FUNCTION "RPA20B_Main" : Void   // FC43, SCL
{ S7_Optimized_Access := 'FALSE' }
VERSION : 0.1
BEGIN


       IF "RPA20B_manual_DOWN" THEN //manual move down
           "RPA20_motor_up" := false;
           "RPA20B_motor_down" := "RPA20B_manual_move";
       ELSIF "RPA20B_manual_UP" THEN // manual move up
           "RPA20_motor_up" := "RPA20B_manual_move";
           "RPA20B_motor_down" := false;
       ELSE // automatic mode operator 1
           "RPA20B_handler_op_1"();
       END_IF;

      "RPA20B_handler_op_2"();

      // blikání LED na tlačítkách

      "RPA20B_open_door_LED_green" := "Clock_0.5Hz" AND ("RPA20B_blend_presence_sensor_1" OR "RPA20B_blend_presence_sensor_2")AND (NOT "RPA20B_open_drawer");

      IF "RPA20B_datablock".RPA20B_station_monitoring_send = true THEN
          "RPA20B_datablock".RPA20B_station_monitoring_send := NOT "pa20b_station_monitoring"(station_activity_state := "RPA20B_ES_feedback",
                                                                                              blend_senzor_l := "RPA20B_blend_presence_sensor_2",
                                                                                              blend_senzor_r := "RPA20B_blend_presence_sensor_1",
                                                                                              server_connection := "tcp_datablock".tcp_connection,
                                                                                              index:="tcp_datablock".<??.?>);
      ELSE
          IF "RPA20B_datablock".RPA20B_activity_state_pre <> "RPA20B_ES_feedback" OR 
              "RPA20B_datablock".RPA20B_left_cover_pressence_sensor_pre <> "RPA20B_blend_presence_sensor_2" OR
              "RPA20B_datablock".RPA20B_right_cover_pressence_sensor_pre <> "RPA20B_blend_presence_sensor_1" THEN
              "RPA20B_datablock".RPA20B_station_monitoring_send := true;
          END_IF;

          "RPA20B_datablock".RPA20B_activity_state_pre := "RPA20B_ES_feedback";
          "RPA20B_datablock".RPA20B_left_cover_pressence_sensor_pre := "RPA20B_blend_presence_sensor_2";
          "RPA20B_datablock".RPA20B_right_cover_pressence_sensor_pre := "RPA20B_blend_presence_sensor_1";
      END_IF;
      IF "RPA20B_manual_UP" THEN
          "RPA20B_Camera_Result_OK" := false;
          "RPA20B_Camera_Result_NOK" := false;
      END_IF;
      "RPA20B_Camera_Trigger" := "RPA20B_Camera_Start_Test";
      "RPA20B_Camera_TrafficLight_Green" := "RPA20B_Camera_Result_OK";
      "RPA20B_Camera_TrafficLight_Red" := "RPA20B_Camera_Result_NOK";
END_FUNCTION

FUNCTION "build_new_record" : Void   // FC44, SCL
{ S7_Optimized_Access := 'FALSE' }
VERSION : 0.1
BEGIN


   #temp_string := CONCAT(IN1 := '$'172', IN2 := "RPA60_DataBlock".RPA60_frame_order);
   #temp_string := CONCAT(IN1 := #temp_string, IN2 := '$', ');
   Strg_TO_Chars(Strg := #temp_string,
                 pChars := 0,
                 Cnt => #i,
                 Chars := #temp_record);

   #chars := 0;
   WHILE #record_in[#chars] <> '?' DO
       #temp_record[#chars+#i] := #record_in[#chars];
      #chars := #chars + 1;
   END_WHILE;

   #temp_record[#chars + #i] := '$L';
   #record_data := #temp_record;

   #i := 0;
   Strg_TO_Chars(Strg:='$'ID$' ,$'frame_code$', $'frame_order$', $'configuration$', $'PA30R_date_time$', $'PA60R_date_time$', ',
                 pChars:=0,
                 Cnt=>#chars,
                 Chars:=#temp_record);

   Strg_TO_Chars(Strg := '$'PA30R_Primer_207_SIKA$', $'PA30R_Remover_208_SIKA$', $'PA30R_rework$', $'PA60R_rework$', $'PA30R_cyclus_completed$', $'PA60R_cyclus_completed$'$L',
                 pChars := #chars,
                 Cnt => #i,
                 Chars := #temp_record);

   #record_items := #temp_record;
END_FUNCTION

FUNCTION "copyAndFill" : Void   // FC45, SCL
{ S7_Optimized_Access := 'FALSE' }
VERSION : 0.1
BEGIN




   //copy the input string to the output string
   #index := 1;
   #inputStringLen := LEN(#stringIn);
   #copyAndFill := '';
   IF #char_number >= #inputStringLen THEN
       WHILE #index <= #char_number DO
           IF #index >= (#char_number - #inputStringLen+1) THEN
               IF #stringIn[#index - (#char_number - #inputStringLen)] <> #charReplace THEN
                   #copyAndFill := CONCAT(IN1 := #copyAndFill, IN2 := #stringIn[#index - (#char_number - #inputStringLen)]);
               ELSE
                   #copyAndFill := CONCAT(IN1 := #copyAndFill, IN2 := #characterFill);
               END_IF;
           ELSE
               #copyAndFill := CONCAT(IN1 := #copyAndFill, IN2 := #characterFill);
           END_IF;

           #index := #index + 1;
       END_WHILE;
   END_IF;
END_FUNCTION

FUNCTION "RPA10B_handler_function" : Void   // FC48, SCL
{ S7_Optimized_Access := 'FALSE' }
VERSION : 0.1
BEGIN
END_FUNCTION

FUNCTION "RPA10B_idler_presence_handler" : Void   // FC49, SCL
{ S7_Optimized_Access := 'FALSE' }
VERSION : 0.1
BEGIN

   (*
   pokud je big fail state odemčený pak se podprogram vykoná

   pokud přítlačné kolečko ve stavu využíváno pak je rozlišováno jestli se jedná o stav ve kterém se čeká na vyjmutí z dokovací stanice a nebo jestli již je vyjmuto z dokovací stanice

   pokud se jedná o stav kdy se čeká na vyjmutí z dokovací stanice musí blikat světelná kontrolka přítlačného kolečka a být nastaven vnitřní stav stanice OK

   pokud se jedná o stav kdy již je přítlačné kolečko z dokovací stanice vyjmuto kontroluje se zda není vloženo zpátky před expirací časovače

   pokud je přítlačné kolečko vloženo do dokovací stanice před expirací časovače dojde k nastavení stavu big fail a blikání světelné kontrolky přítlačného kolečka

   *)

   IF (#bigFailStateLock = 0 OR #bigFailStateLock = #bigFailStateIdentifire OR #bigFailStateLock = #bigFailStateIdentifire + 100) AND
       #errorStateLock = 0 AND
       #fatalErrorStateLock = 0 THEN

       //blikání a svícení světelné kontrolky přítlačného kolečka
       //#bottlePresenceSensor AND "Clock_0.5Hz" AND #bottleInUsage
      // #rollerLED := (NOT #rollerPresenceSensor) OR (#rollerPresenceSensor AND "Clock_0.5Hz" AND #roller_in_use);
       //#rollerLED := (NOT #rollerPresenceSensor) OR (#rollerPresenceSensor AND #rollerUsageInterval[#workCyclusControlVariable] AND "Clock_0.5Hz");

       IF #bigFailStateLock = #bigFailStateIdentifire  THEN
           "setOKState"(confirm := true,
                        identifier := #bigFailStateIdentifire,
                        confirm_blinking := false,
                        blinkConfirmButton => #confirmButtonLed,
                        stateLock := #bigFailStateLock);
       ELSIF #bigFailStateLock = #bigFailStateIdentifire+100 AND #idler_presence_sensor = true THEN
               "setOKState"(confirm := #confirmButton,
                            identifier := #bigFailStateIdentifire+100,
                            confirm_blinking := true,
                            blinkConfirmButton => #confirmButtonLed,
                            stateLock := #bigFailStateLock);
       END_IF;
       //kontrola přítomnosti kolečka v pracovním cyklu
       IF #idler_in_use THEN
           "RPA10B_datablock".RPA10B_idler_checking_dalay := false;
           //nekontroluje první stav a poslední stav ve kterém je přítlačné kolečko používáno -> stav ve kterém se mění mění přítomnost kolečka v dokovací stanici
               IF #idler_presence_sensor THEN
                   IF #idler_taking THEN
                       IF "setBigFailState"(identifier := #bigFailStateIdentifire,
                                                error_state_lock:="RPA10B_datablock".PA10B_error_state_lock, fatal_state_error:="RPA10B_datablock".PA10B_fatal_error_state_lock, badfailStateLock := #bigFailStateLock) THEN
                           ;
                       END_IF;
                   END_IF;
               END_IF;
        ELSE
            IF (NOT #idler_presence_sensor) THEN
                IF "RPA10B_datablock".RPA10B_idler_checking_dalay THEN
                    IF "setBigFailState"(identifier := #bigFailStateIdentifire + 100,
                                             error_state_lock := "RPA10B_datablock".PA10B_error_state_lock, fatal_state_error := "RPA10B_datablock".PA10B_fatal_error_state_lock, badfailStateLock := #bigFailStateLock) THEN
                        ;
                    END_IF;
                ELSE
                    "RPA10B_datablock".RPA10B_idler_checking_dalay := "Clock_0.5Hz";
                END_IF;
            END_IF;
       END_IF;
   END_IF;
END_FUNCTION

FUNCTION "server_connection_handler" : Void   // FC50, SCL
{ S7_Optimized_Access := 'FALSE' }
VERSION : 0.1
BEGIN
   IF #database_connection = true THEN
       IF #error_state_lock = #error_state_lock_identifier THEN
           #error_state_lock := 0;
       END_IF;
   ELSE
       IF #fatal_error_state_lock = 0 AND #error_state_lock = 0 THEN
           #error_state_lock := #error_state_lock_identifier;
       END_IF;
   END_IF;
END_FUNCTION

FUNCTION "station_reset" : Void   // FC51, SCL
{ S7_Optimized_Access := 'FALSE' }
VERSION : 0.1
BEGIN
   #index := 1;

   WHILE (#index < 6) DO
       #fs_funel_control[#index] := false;
       #fs_show_fill_button[#index] := false;
       #index := #index + 1;
   END_WHILE;

   #funel_1 := false;
   #funel_2 := false;
   #funel_3 := false;
   #funel_4 := false;
   #funel_5 := false;

   #fs_chemical_type := 0;
   #hmi_label_index := 0;


   #fill_bottle_step := 9;
   #shake_deinit := true;
   #print_sp_bottle_label_step := 8;



   #fs_show_manual_or_scan := false;
   #fs_show_button := false;
   #fs_reset_e := false;
END_FUNCTION

FUNCTION "time_compare" : Void   // FC52, LAD
{ S7_Optimized_Access := 'FALSE' }
VERSION : 0.1
BEGIN

REGION Network 1
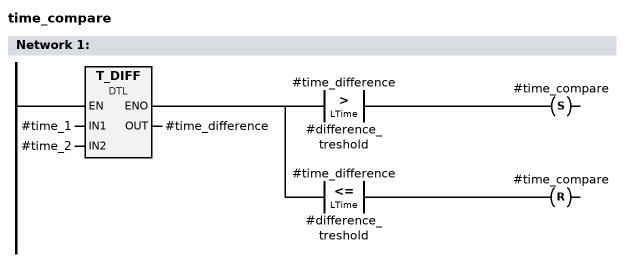
   // ENO of a box is taken as its EN; it also drops when the box reports an error
   #time_difference := T_DIFF(IN1 := #time_1, IN2 := #time_2);
   IF #time_difference > #difference_treshold THEN #time_compare := TRUE; END_IF;
   IF #time_difference <= #difference_treshold THEN #time_compare := FALSE; END_IF;
END_REGION
END_FUNCTION

FUNCTION "RPA30_Handler_function_A" : Void   // FC53, SCL
{ S7_Optimized_Access := 'FALSE' }
VERSION : 0.1
BEGIN
END_FUNCTION

FUNCTION "pa10r_station_monitoring" : Void   // FC54, SCL
{ S7_Optimized_Access := 'FALSE' }
VERSION : 0.1
BEGIN
   #pa10r_station_monitoring := false;
   (*
   IF #server_connection = true THEN
       IF "send_msg_to_pc_DB".DONE THEN
           "rcv_msg_from_pc_DB"(size := 1024,
                                time_out_interval := #lock);

           IF "rcv_msg_from_pc_DB".time_out = true THEN
               "send_msg_to_pc_DB".DONE := false;
               "rcv_msg_from_pc_DB".DONE := false;
               #server_connection := false;
           END_IF;

           IF "rcv_msg_from_pc_DB".DONE THEN
               "send_msg_to_pc_DB".DONE := false;
               "rcv_msg_from_pc_DB".DONE := false;
               "send_msg_to_pc_DB".synchronization := 0;
               "rcv_msg_from_pc_DB".synchronization := 0;
               #server_connection := true;
               #pa10r_station_monitoring := true;
           END_IF;
       ELSE

           //command 
           Strg_TO_Chars(Strg := 'PA10R_STATE~',
                         pChars := 0,
                         Cnt => #chars,
                         Chars := #chars_out);
           #i := #chars;

           // station state 
           IF #station_activity_state = true THEN
               IF #fatal_error_state > 0 THEN
                   CASE #fatal_error_state OF
                       150:
                           Strg_TO_Chars(Strg := '<html>Station state: Y axis<br>valve lock error</html>~',
                                         pChars := #i,
                                         Cnt => #chars,
                                         Chars := #chars_out);
                       160:
                           Strg_TO_Chars(Strg := '<html>Station state: X axis<br>valve lock error</html>~',
                                         pChars := #i,
                                         Cnt => #chars,
                                         Chars := #chars_out);
                       ELSE
                           Strg_TO_Chars(Strg := 'Station state: Unknown~',
                                         pChars := #i,
                                         Cnt => #chars,
                                         Chars := #chars_out);
                   END_CASE;
               ELSE
                   IF #error_state > 0 THEN
                       Strg_TO_Chars(Strg := 'Station state: Unknown~',
                                     pChars := #i,
                                     Cnt => #chars,
                                     Chars := #chars_out);
                   ELSE
                       IF #big_fail_state > 0 THEN
                           Strg_TO_Chars(Strg := 'Station state: Unknown~',
                                         pChars := #i,
                                         Cnt => #chars,
                                         Chars := #chars_out);
                       ELSE
                           IF #fail_state > 0 THEN
                               CASE #fail_state OF
                                   110:
                                       Strg_TO_Chars(Strg := 'Station state: Felt box is empty~',
                                                     pChars := #i,
                                                     Cnt => #chars,
                                                     Chars := #chars_out);
                                   200:  // Statement section case 2 to 4
                                       Strg_TO_Chars(Strg := '<html>Station state: Primer DV594V1<br>in primer box</html>~',
                                                     pChars := #i,
                                                     Cnt => #chars,
                                                     Chars := #chars_out);
                                   201:
                                       Strg_TO_Chars(Strg := '<html>Station state: Activator DW646<br>in primer box</html>~',
                                                     pChars := #i,
                                                     Cnt => #chars,
                                                     Chars := #chars_out);
                                   202:
                                       Strg_TO_Chars(Strg := '<html>Station state: Primer 207<br>in primer box</html>~',
                                                     pChars := #i,
                                                     Cnt => #chars,
                                                     Chars := #chars_out);
                                   300:
                                       Strg_TO_Chars(Strg := '<html>Station state: Primer DV594V1<br>out of primer box</html>~',
                                                     pChars := #i,
                                                     Cnt => #chars,
                                                     Chars := #chars_out);
                                   301:
                                       Strg_TO_Chars(Strg := '<html>Station state: Activator DW646<br>out of primer box</html>~',
                                                     pChars := #i,
                                                     Cnt => #chars,
                                                     Chars := #chars_out);
                                   302:
                                       Strg_TO_Chars(Strg := '<html>Station state: Primer 207<br>out of primer box</html>~',
                                                     pChars := #i,
                                                     Cnt => #chars,
                                                     Chars := #chars_out);
                                   303:
                                       Strg_TO_Chars(Strg := '<html>Station state: Remover 208<br>out of primer box</html>~',
                                                     pChars := #i,
                                                     Cnt => #chars,
                                                     Chars := #chars_out);
                                   6:
                                       Strg_TO_Chars(Strg := 'Station state: Remover 208 expired~',
                                                     pChars := #i,
                                                     Cnt => #chars,
                                                     Chars := #chars_out);
                                   ELSE  // Statement section ELSE
                                       Strg_TO_Chars(Strg := 'Station state: Unknown~',
                                                     pChars := #i,
                                                     Cnt => #chars,
                                                     Chars := #chars_out);
                               END_CASE;

                           ELSE
                               Strg_TO_Chars(Strg := 'Station state: OK~',
                                             pChars := #i,
                                             Cnt => #chars,
                                             Chars := #chars_out);
                           END_IF;
                       END_IF;
                   END_IF;
               END_IF;
           ELSE
               Strg_TO_Chars(Strg := 'Station state: Inactive~',
                             pChars := #i,
                             Cnt => #chars,
                             Chars := #chars_out);
           END_IF;

           #i := #i+#chars;

           // work cyclus state 

           IF #work_cyclus_state = "RPA10R_hmi_go_to_home_position" THEN
               Strg_TO_Chars(Strg := 'Work cyclus state: Waiting for home position~',
                             pChars := #i,
                             Cnt => #chars,
                             Chars := #chars_out);
           ELSIF #work_cyclus_state = "RPA10R_hmi_scan_frame" THEN
               Strg_TO_Chars(Strg := 'Work cyclus state: Scan frame~',
                             pChars := #i,
                             Cnt => #chars,
                             Chars := #chars_out);
           ELSIF #work_cyclus_state = "RPA10R_hmi_take_bottle_1" THEN
               Strg_TO_Chars(Strg := 'Work cyclus state: Take activator DW 646~',
                             pChars := #i,
                             Cnt => #chars,
                             Chars := #chars_out);
           ELSIF #work_cyclus_state = "RPA10R_hmi_scan_bottle" THEN
               Strg_TO_Chars(Strg := 'Work cyclus state: Scan bottle~',
                             pChars := #i,
                             Cnt => #chars,
                             Chars := #chars_out);
           ELSIF #work_cyclus_state = "RPA10R_hmi_change_pad" THEN
               Strg_TO_Chars(Strg := 'Work cyclus state: Change pad~',
                             pChars := #i,
                             Cnt => #chars,
                             Chars := #chars_out);
           ELSIF #work_cyclus_state = "RPA10R_hmi_apply_bottle_1_on_side_5_5" OR #work_cyclus_state = "RPA10R_hmi_apply_bottle_1_on_side_5" THEN
               Strg_TO_Chars(Strg := 'Work cyclus state: Apply activator on frame~',
                             pChars := #i,
                             Cnt => #chars,
                             Chars := #chars_out);
           ELSIF #work_cyclus_state = "RPA10R_hmi_turn_clockwise" THEN
               Strg_TO_Chars(Strg := 'Work cyclus state: Turn frame clockwise~',
                             pChars := #i,
                             Cnt => #chars,
                             Chars := #chars_out);
           ELSIF #work_cyclus_state = "RPA10R_hmi_take_bottle_2" THEN
               Strg_TO_Chars(Strg := 'Work cyclus state: Take bottle of primer DV954~',
                             pChars := #i,
                             Cnt => #chars,
                             Chars := #chars_out);
           ELSIF #work_cyclus_state = "RPA10R_hmi_whipe_off_side_5_5" OR #work_cyclus_state = "RPA10R_hmi_whipe_off_side_5" THEN
               Strg_TO_Chars(Strg := '<html>Work cyclus state: Wipe off activator<br> from frame</html>~',
                             pChars := #i,
                             Cnt => #chars,
                             Chars := #chars_out);
           ELSIF #work_cyclus_state = "RPA10R_hmi_apply_bottle_2_on_side_5_5" OR #work_cyclus_state = "RPA10R_hmi_apply_bottle_2_on_side_5" THEN
               Strg_TO_Chars(Strg := 'Work cyclus state: Apply primer on frame~',
                             pChars := #i,
                             Cnt => #chars,
                             Chars := #chars_out);
           ELSIF #work_cyclus_state = "RPA10R_hmi_put_back_bottle_1" THEN
               Strg_TO_Chars(Strg := '<html>Work cyclus state: Put activator DW 646<br>bottle to primer bar</html>~',
                             pChars := #i,
                             Cnt => #chars,
                             Chars := #chars_out);
           ELSIF #work_cyclus_state = "RPA10R_hmi_put_back_bottle_2" THEN
               Strg_TO_Chars(Strg := '<html>Work cyclus state: Put primer DV954 bottle<br>to primer bar</html>~',
                             pChars := #i,
                             Cnt => #chars,
                             Chars := #chars_out);
           ELSIF #work_cyclus_state = "RPA10R_hmi_take_felt" THEN
               Strg_TO_Chars(Strg := 'Work cyclus state: Take felt~',
                             pChars := #i,
                             Cnt => #chars,
                             Chars := #chars_out);
           ELSIF #work_cyclus_state = "RPA10R_hmi_turn_horizontaly" THEN
               Strg_TO_Chars(Strg := 'Work cyclus state: Turn frame horizontaly~',
                             pChars := #i,
                             Cnt => #chars,
                             Chars := #chars_out);
           ELSIF #work_cyclus_state = "RPA10R_hmi_on_felt_apply_remover" THEN
               Strg_TO_Chars(Strg := 'Work cyclus state: On felt apply remover~',
                             pChars := #i,
                             Cnt => #chars,
                             Chars := #chars_out);
           ELSIF #work_cyclus_state = "RPA10R_hmi_apply_remover_to_side_5" THEN
               Strg_TO_Chars(Strg := 'Work cyclus state: Apply remover 208 on frame~',
                             pChars := #i,
                             Cnt => #chars,
                             Chars := #chars_out);
           ELSIF #work_cyclus_state = "RPA10R_hmi_turn_counterclockwise" THEN
               Strg_TO_Chars(Strg := 'Work cyclus state: Turn frame counterclockwise~',
                             pChars := #i,
                             Cnt => #chars,
                             Chars := #chars_out);
           ELSIF #work_cyclus_state = "RPA10R_hmi_take_bottle_3" THEN
               Strg_TO_Chars(Strg := 'Work cyclus state: Take bottle of primer 207~',
                             pChars := #i,
                             Cnt => #chars,
                             Chars := #chars_out);
           ELSIF #work_cyclus_state = "RPA10R_hmi_put_back_bottle_3" THEN
               Strg_TO_Chars(Strg := '<html>Work cyclus state: Put primer 207 bottle <br> to primer bar</html>~',
                             pChars := #i,
                             Cnt => #chars,
                             Chars := #chars_out);
           ELSIF #work_cyclus_state = "RPA10R_hmi_end_of_cyclus" THEN
               Strg_TO_Chars(Strg := 'Work cyclus state: End of work cyclus~',
                             pChars := #i,
                             Cnt => #chars,
                             Chars := #chars_out);
           ELSIF #work_cyclus_state = 254 THEN
               Strg_TO_Chars(Strg := 'Work cyclus state: Manual mode~',
                             pChars := #i,
                             Cnt => #chars,
                             Chars := #chars_out);
           ELSE
               Strg_TO_Chars(Strg := 'Work cyclus state: Unknown~',
                             pChars := #i,
                             Cnt => #chars,
                             Chars := #chars_out);
           END_IF;

           #i := #i+#chars;
           // home position 
           IF #position_sensor_y AND #position_sensor_x THEN
               Strg_TO_Chars(Strg := 'Home position: Yes~',
                             pChars := #i,
                             Cnt => #chars,
                             Chars := #chars_out);
           ELSE
               Strg_TO_Chars(Strg := 'Home position: No~',
                             pChars := #i,
                             Cnt => #chars,
                             Chars := #chars_out);
           END_IF;

           #i := #i + #chars;
           // current frame code
           Strg_TO_Chars(Strg := 'Current frame code: ',
                         pChars := #i,
                         Cnt => #chars,
                         Chars := #chars_out);
           #i := #i + #chars;
           IF #current_frame_code <> '' THEN
               Strg_TO_Chars(Strg := #current_frame_code,
                             pChars := #i,
                             Cnt => #chars,
                             Chars := #chars_out);
           ELSE
               Strg_TO_Chars(Strg := 'None',
                             pChars := #i,
                             Cnt => #chars,
                             Chars := #chars_out);
           END_IF;
           #i := #i + #chars;

           // station configuration
           IF #station_configuration = 0 THEN
               Strg_TO_Chars(Strg := '~Station configuration: 581A~',
                             pChars := #i,
                             Cnt => #chars,
                             Chars := #chars_out);
           ELSIF #station_configuration = 1 THEN
               Strg_TO_Chars(Strg := '~Station configuration: 581B~',
                             pChars := #i,
                             Cnt => #chars,
                             Chars := #chars_out);
           ELSIF #station_configuration = 2 THEN
               Strg_TO_Chars(Strg := '~Station configuration: 582A~',
                             pChars := #i,
                             Cnt => #chars,
                             Chars := #chars_out);
           ELSIF #station_configuration = 3 THEN
               Strg_TO_Chars(Strg := '~Station configuration: 582B~',
                             pChars := #i,
                             Cnt => #chars,
                             Chars := #chars_out);
           END_IF;

           #i := #i + #chars;

           "send_msg_to_pc_DB"(lock := #chars_out,
                               lock := 1024,
                               time_out_interval := #i,
                               time_out_interval := #lock);
           IF "send_msg_to_pc_DB".time_out = true THEN
               #server_connection := false;
           END_IF;
       END_IF;
   END_IF;
   *)
END_FUNCTION

FUNCTION "pa50r_station_monitoring" : Void   // FC55, SCL
{ S7_Optimized_Access := 'FALSE' }
VERSION : 0.1
BEGIN
   #pa50r_station_monitoring := false;
   (*
   IF #server_connection = true THEN
       IF "send_msg_to_pc_DB".DONE THEN
           "rcv_msg_from_pc_DB"(size := 1024,
                                time_out_interval := #lock);

           IF "rcv_msg_from_pc_DB".time_out = true THEN
               "send_msg_to_pc_DB".DONE := false;
               "rcv_msg_from_pc_DB".DONE := false;
               #server_connection := false;
           END_IF;

           IF "rcv_msg_from_pc_DB".DONE THEN
               "send_msg_to_pc_DB".DONE := false;
               "rcv_msg_from_pc_DB".DONE := false;
               "send_msg_to_pc_DB".synchronization := 0;
               "rcv_msg_from_pc_DB".synchronization := 0;
               #server_connection := true;
               #pa50r_station_monitoring := true;
           END_IF;
       ELSE

           //command 
           Strg_TO_Chars(Strg := 'PA50R_STATE~',
                         pChars := 0,
                         Cnt => #chars,
                         Chars := #chars_out);
           #i := #chars;

           //station state
           IF #station_activity_state = true THEN
               IF #fatal_error_state > 0 THEN
                   Strg_TO_Chars(Strg := 'Station state: Unknown~',
                                 pChars := #i,
                                 Cnt => #chars,
                                 Chars := #chars_out);
               ELSE
                   IF #error_state > 0 THEN
                       CASE #error_state OF
                           21000:
                               Strg_TO_Chars(Strg := 'Station state: Frame already processed~',
                                             pChars := #i,
                                             Cnt => #chars,
                                             Chars := #chars_out);
                           22000:
                               Strg_TO_Chars(Strg := 'Station state:Frame was not on previous station~',
                                             pChars := #i,
                                             Cnt => #chars,
                                             Chars := #chars_out);
                           23000:
                               Strg_TO_Chars(Strg := 'Station state: Frame has more then 8 hours~',
                                             pChars := #i,
                                             Cnt => #chars,
                                             Chars := #chars_out);
                           24000:
                               Strg_TO_Chars(Strg := 'Station state: Frame has less then 10 minutes~',
                                             pChars := #i,
                                             Cnt => #chars,
                                             Chars := #chars_out);
                           25000:
                               Strg_TO_Chars(Strg := 'Station state: Frame is not in database~',
                                             pChars := #i,
                                             Cnt => #chars,
                                             Chars := #chars_out);
                           26000:
                               Strg_TO_Chars(Strg := 'Station state: Bad station configuration~',
                                             pChars := #i,
                                             Cnt => #chars,
                                             Chars := #chars_out);
                           ELSE  // Statement section ELSE
                               Strg_TO_Chars(Strg := 'Station state: Unknown~',
                                             pChars := #i,
                                             Cnt => #chars,
                                             Chars := #chars_out);
                       END_CASE;

                       Strg_TO_Chars(Strg := 'Station state: Unknown~',
                                     pChars := #i,
                                     Cnt => #chars,
                                     Chars := #chars_out);
                   ELSE
                       IF #big_fail_state > 0 THEN
                           Strg_TO_Chars(Strg := 'Station state: Unknown~',
                                         pChars := #i,
                                         Cnt => #chars,
                                         Chars := #chars_out);
                       ELSE
                           IF #fail_state > 0 THEN
                                       Strg_TO_Chars(Strg := 'Station state: Unknown~',
                                                     pChars := #i,
                                                     Cnt => #chars,
                                                     Chars := #chars_out);
                           ELSE
                               Strg_TO_Chars(Strg := 'Station state: OK~',
                                             pChars := #i,
                                             Cnt => #chars,
                                             Chars := #chars_out);
                           END_IF;
                       END_IF;
                   END_IF;
               END_IF;
           ELSE
               Strg_TO_Chars(Strg := 'Station state: Inactive~',
                             pChars := #i,
                             Cnt => #chars,
                             Chars := #chars_out);
           END_IF;

           #i := #i+#chars;

           //work cyclus state

           IF #work_cyclus_state = "RPA50_hmi_go_to_home_position" THEN
               Strg_TO_Chars(Strg := 'Work cyclus state: Waiting for home position~',
                             pChars := #i,
                             Cnt => #chars,
                             Chars := #chars_out);
           ELSIF #work_cyclus_state = "RPA50_hmi_scan_frame" THEN
               Strg_TO_Chars(Strg := 'Work cyclus state: Scan frame code~',
                             pChars := #i,
                             Cnt => #chars,
                             Chars := #chars_out);
           ELSIF #work_cyclus_state = "RPA50_hmi_apply_tape" THEN
               Strg_TO_Chars(Strg := '<html>Work cyclus state: Application of tape <br>on every sides of grame</hmt>~',
                             pChars := #i,
                             Cnt => #chars,
                             Chars := #chars_out);
           ELSIF #work_cyclus_state = "RPA50_hmi_end_of_cyclus" THEN
               Strg_TO_Chars(Strg := 'Work cyclus state: End of work cyclus~',
                             pChars := #i,
                             Cnt => #chars,
                             Chars := #chars_out);
           ELSE
               Strg_TO_Chars(Strg := 'Work cyclus state: Unknown~',
                             pChars := #i,
                             Cnt => #chars,
                             Chars := #chars_out);
           END_IF;

           #i := #i+#chars;
           //home position
           IF #position_sensor_y THEN
               Strg_TO_Chars(Strg := 'Home position: Yes~',
                             pChars := #i,
                             Cnt => #chars,
                             Chars := #chars_out);
           ELSE
               Strg_TO_Chars(Strg := 'Home position: No~',
                             pChars := #i,
                             Cnt => #chars,
                             Chars := #chars_out);
           END_IF;

           #i := #i + #chars;
           //current frame code
           Strg_TO_Chars(Strg := 'Current frame code: ',
                         pChars := #i,
                         Cnt => #chars,
                         Chars := #chars_out);
           #i := #i + #chars;
           IF #current_frame_code <> '' THEN
               Strg_TO_Chars(Strg := #current_frame_code,
                             pChars := #i,
                             Cnt => #chars,
                             Chars := #chars_out);
           ELSE
               Strg_TO_Chars(Strg := 'None',
                             pChars := #i,
                             Cnt => #chars,
                             Chars := #chars_out);
           END_IF;
           #i := #i + #chars;

           //station configuration
           IF #station_configuration = 0 THEN
               Strg_TO_Chars(Strg := '~Station configuration: 581A',
                             pChars := #i,
                             Cnt => #chars,
                             Chars := #chars_out);
           ELSIF #station_configuration = 1 THEN
               Strg_TO_Chars(Strg := '~Station configuration: 581B',
                             pChars := #i,
                             Cnt => #chars,
                             Chars := #chars_out);
           ELSIF #station_configuration = 2 THEN
               Strg_TO_Chars(Strg := '~Station configuration: 582A',
                             pChars := #i,
                             Cnt => #chars,
                             Chars := #chars_out);
           ELSIF #station_configuration = 3 THEN
               Strg_TO_Chars(Strg := '~Station configuration: 582B',
                             pChars := #i,
                             Cnt => #chars,
                             Chars := #chars_out);
           END_IF;

           #i := #i + #chars;

           "send_msg_to_pc_DB"(time_out_interval := #chars_out,
                               time_out_interval := 1024,
                               lock := #i,
                               lock := #lock);
           IF "send_msg_to_pc_DB".time_out = true THEN
               #server_connection := false;
           END_IF;
       END_IF;
   END_IF;
   *)
END_FUNCTION

FUNCTION "pa60r_station_monitoring" : Void   // FC56, SCL
{ S7_Optimized_Access := 'FALSE' }
VERSION : 0.1
BEGIN
   #pa60r_station_monitoring := false;
   IF #server_connection = true THEN
       IF #index = 255 THEN
       (* command *)
           Strg_TO_Chars(Strg := 'PA60R_STATE~',
                         pChars := 0,
                         Cnt => #chars,
                         Chars := #temp_buffer);
           #i := #chars;

           (* station state *)
           IF #station_activity_state = true THEN
               IF #fatal_error_state > 0 THEN
                   CASE #fatal_error_state OF
                       150:  // Statement section case 1
                           Strg_TO_Chars(Strg := 'Station state: Y axis valve lock error~',
                                         pChars := #i,
                                         Cnt => #chars,
                                         Chars := #temp_buffer);
                       170:
                           Strg_TO_Chars(Strg := 'Station state: Bad frame code~',
                                         pChars := #i,
                                         Cnt => #chars,
                                         Chars := #temp_buffer);
                       180:
                           Strg_TO_Chars(Strg := 'Station state: Bad hardware configuration~',
                                         pChars := #i,
                                         Cnt => #chars,
                                         Chars := #temp_buffer);
                       230:
                           Strg_TO_Chars(Strg := 'Station state: Seal presence error~',
                                         pChars := #i,
                                         Cnt => #chars,
                                         Chars := #temp_buffer);
                       293:
                           Strg_TO_Chars(Strg := 'Station state: Change sealing fixtures~',
                                         pChars := #i,
                                         Cnt => #chars,
                                         Chars := #temp_buffer);
                       ELSE  // Statement section ELSE
                           Strg_TO_Chars(Strg := 'Station state: Unknown~',
                                         pChars := #i,
                                         Cnt => #chars,
                                         Chars := #temp_buffer);
                   END_CASE;
               ELSE
                   IF #error_state > 0 THEN
                       CASE #error_state OF
                           20000:
                               Strg_TO_Chars(Strg := 'Station state: Frame already processed~',
                                             pChars := #i,
                                             Cnt => #chars,
                                             Chars := #temp_buffer);
                           21000:
                               Strg_TO_Chars(Strg := 'Station state:Frame was not on previous station~',
                                             pChars := #i,
                                             Cnt => #chars,
                                             Chars := #temp_buffer);
                           23000:
                               Strg_TO_Chars(Strg := 'Station state: Frame has more then 8 hours~',
                                             pChars := #i,
                                             Cnt => #chars,
                                             Chars := #temp_buffer);
                           24000:
                               Strg_TO_Chars(Strg := 'Station state: Frame has less then 10 minutes~',
                                             pChars := #i,
                                             Cnt => #chars,
                                             Chars := #temp_buffer);
                           25000:
                               Strg_TO_Chars(Strg := 'Station state: Frame is not in database~',
                                             pChars := #i,
                                             Cnt => #chars,
                                             Chars := #temp_buffer);
                           26000:
                               Strg_TO_Chars(Strg := 'Station state: Bad station configuration~',
                                             pChars := #i,
                                             Cnt => #chars,
                                             Chars := #temp_buffer);
                           ELSE  // Statement section ELSE
                               Strg_TO_Chars(Strg := 'Station state: Unknown~',
                                             pChars := #i,
                                             Cnt => #chars,
                                             Chars := #temp_buffer);
                       END_CASE;

                       Strg_TO_Chars(Strg := 'Station state: Unknown~',
                                     pChars := #i,
                                     Cnt => #chars,
                                     Chars := #temp_buffer);
                   ELSE
                       IF #big_fail_state > 0 THEN
                           CASE #big_fail_state OF
                               120:  // Statement section case 1
                                   Strg_TO_Chars(Strg := 'Station state: Roller out of home position~',
                                                 pChars := #i,
                                                 Cnt => #chars,
                                                 Chars := #temp_buffer);

                               ELSE
                                   Strg_TO_Chars(Strg := 'Station state: Unknown~',
                                                 pChars := #i,
                                                 Cnt => #chars,
                                                 Chars := #temp_buffer);
                           END_CASE;


                       ELSE
                           IF #fail_state > 0 THEN
                               Strg_TO_Chars(Strg := 'Station state: Unknown~',
                                             pChars := #i,
                                             Cnt => #chars,
                                             Chars := #temp_buffer);
                           ELSE
                               Strg_TO_Chars(Strg := 'Station state: OK~',
                                             pChars := #i,
                                             Cnt => #chars,
                                             Chars := #temp_buffer);
                           END_IF;
                       END_IF;
                   END_IF;
               END_IF;
           ELSE
               Strg_TO_Chars(Strg := 'Station state: Inactive~',
                             pChars := #i,
                             Cnt => #chars,
                             Chars := #temp_buffer);
           END_IF;

           #i := #i + #chars;

           (* work cyclus state *)

           IF #work_cyclus_state = "RPA60_hmi_go_to_home_position" THEN
               Strg_TO_Chars(Strg := 'Work cyclus state: Waiting for home position~',
                             pChars := #i,
                             Cnt => #chars,
                             Chars := #temp_buffer);
           ELSIF #work_cyclus_state = "RPA60_hmi_scan_frame" THEN
               Strg_TO_Chars(Strg := 'Work cyclus state: Scan frame code~',
                             pChars := #i,
                             Cnt => #chars,
                             Chars := #temp_buffer);
           ELSIF #work_cyclus_state = "RPA60_hmi_turn_frame_clockwise" THEN
               Strg_TO_Chars(Strg := 'Work cyclus state: Turn frame clockwise~',
                             pChars := #i,
                             Cnt => #chars,
                             Chars := #temp_buffer);
           ELSIF #work_cyclus_state = "RPA60_hmi_put_sealing_in_the_ficture" THEN
               Strg_TO_Chars(Strg := '<html>Work cyclus state: Put sealing in the fixture<br>and glue sealing on the desk</html>~',
                             pChars := #i,
                             Cnt => #chars,
                             Chars := #temp_buffer);
           ELSIF #work_cyclus_state = "RPA60_hmi_press_sealing_with_roller" THEN
               Strg_TO_Chars(Strg := 'Work cyclus state: Press sealing with roller~',
                             pChars := #i,
                             Cnt => #chars,
                             Chars := #temp_buffer);
           ELSIF #work_cyclus_state = "RPA60_hmi_put_roller_to_home_position" THEN
               Strg_TO_Chars(Strg := 'Work cyclus state: Put roller to home position~',
                             pChars := #i,
                             Cnt => #chars,
                             Chars := #temp_buffer);
           ELSIF #work_cyclus_state = "RPA60_hmi_seals_pressence_testing" THEN
               Strg_TO_Chars(Strg := 'Work cyclus state: Seals pressence testing~',
                             pChars := #i,
                             Cnt => #chars,
                             Chars := #temp_buffer);
           ELSIF #work_cyclus_state = "RPA60_hmi_seals_missing" THEN
               Strg_TO_Chars(Strg := 'Work cyclus state: Seals missing on the frame~',
                             pChars := #i,
                             Cnt => #chars,
                             Chars := #temp_buffer);
           ELSIF #work_cyclus_state = "RPA60_hmi_scan_printed_label" THEN
               Strg_TO_Chars(Strg := 'Work cyclus state: Scan printed label~',
                             pChars := #i,
                             Cnt => #chars,
                             Chars := #temp_buffer);
           ELSIF #work_cyclus_state = "RPA60_hmi_label_is_wrong" THEN
               Strg_TO_Chars(Strg := 'Work cyclus state: Scanned label is wrong~',
                             pChars := #i,
                             Cnt => #chars,
                             Chars := #temp_buffer);
           ELSIF #work_cyclus_state = "RPA60_hmi_cyclus_finished_ok" THEN
               Strg_TO_Chars(Strg := 'Work cyclus state: Work cyclus finished OK~',
                             pChars := #i,
                             Cnt => #chars,
                             Chars := #temp_buffer);
           ELSIF #work_cyclus_state = "RPA60_hmi_check_agin" THEN
               Strg_TO_Chars(Strg := 'Work cyclus state: Check sealing agin~',
                             pChars := #i,
                             Cnt => #chars,
                             Chars := #temp_buffer);
           ELSE
               Strg_TO_Chars(Strg := 'Work cyclus state: Unknown~',
                             pChars := #i,
                             Cnt => #chars,
                             Chars := #temp_buffer);
           END_IF;

           #i := #i + #chars;
           (* home position *)
           IF #position_sensor_y THEN
               Strg_TO_Chars(Strg := 'Home position: Yes~',
                             pChars := #i,
                             Cnt => #chars,
                             Chars := #temp_buffer);
           ELSE
               Strg_TO_Chars(Strg := 'Home position: No~',
                             pChars := #i,
                             Cnt => #chars,
                             Chars := #temp_buffer);
           END_IF;

           #i := #i + #chars;
           (* current frame code *)
           Strg_TO_Chars(Strg := 'Current frame code: ',
                         pChars := #i,
                         Cnt => #chars,
                         Chars := #temp_buffer);
           #i := #i + #chars;
           IF #current_frame_code <> '' THEN
               Strg_TO_Chars(Strg := #current_frame_code,
                             pChars := #i,
                             Cnt => #chars,
                             Chars := #temp_buffer);
           ELSE
               Strg_TO_Chars(Strg := 'None',
                             pChars := #i,
                             Cnt => #chars,
                             Chars := #temp_buffer);
           END_IF;
           #i := #i + #chars;

           (* station configuration *)
           IF #station_configuration = 0 THEN
               Strg_TO_Chars(Strg := '~Station configuration: 581A~',
                             pChars := #i,
                             Cnt => #chars,
                             Chars := #temp_buffer);
           ELSIF #station_configuration = 1 THEN
               Strg_TO_Chars(Strg := '~Station configuration: 581B~',
                             pChars := #i,
                             Cnt => #chars,
                             Chars := #temp_buffer);
           ELSIF #station_configuration = 2 THEN
               Strg_TO_Chars(Strg := '~Station configuration: 582A~',
                             pChars := #i,
                             Cnt => #chars,
                             Chars := #temp_buffer);
           ELSIF #station_configuration = 3 THEN
               Strg_TO_Chars(Strg := '~Station configuration: 582B~',
                             pChars := #i,
                             Cnt => #chars,
                             Chars := #temp_buffer);
           END_IF;

           #i := #i + #chars;
           #temp_buffer[#i] :='$L';
           #msg_index := "tcp_send"(#temp_buffer);
           IF #msg_index <> 255 THEN
               #index := #msg_index;
           END_IF;
       ELSE
           IF "tcp_rcv"(msg_index := #index, rcv_data => #temp_buffer) = true THEN
               #index := 255;
               #pa60r_station_monitoring := true;
           END_IF;
       END_IF;
   END_IF;
END_FUNCTION

FUNCTION "parse_input_data" : Void   // FC57, SCL
{ S7_Optimized_Access := 'FALSE' }
VERSION : 0.1
BEGIN
   #index := 0;
   #parse_input_data := '';
   WHILE #String_in[#index] <> '$00' AND #String_in[#index] <> '?' AND #index <= 255 DO
       #parse_input_data := CONCAT(IN1 := #parse_input_data, IN2 := #String_in[#index]);
       #index := #index + 1;
   END_WHILE;
END_FUNCTION

FUNCTION "sub_string" : Void   // FC58, SCL
{ S7_Optimized_Access := 'FALSE' }
VERSION : 0.1
BEGIN